       #tempInternalError := MOVE_BLK_VARIANT(SRC := #initialValue,
                                              COUNT := 1,
                                              SRC_INDEX := 0,
                                              DEST_INDEX := #tempSizeCounter,
                                              DEST => #buffer);
     END_FOR;
     IF (#tempInternalError <> #NO_INTERNAL_ERROR) THEN
       #error := true;
       #statusID := #ERROR_MOVE_BLK_VARIANT;
       #status := INT_TO_WORD(#tempInternalError);
     END_IF;
     RETURN;
   END_IF;

   //-----------Program code execution, depending on the Mode parameter-------------
   // The execution of the instructions depends on the signal state of the Mode parameter.

   IF #mode = #NEXT_TASK_TO_EXECUTE THEN


     // If the Mode parameter has the signal state "0",
     // the first entry from the passed ring buffer is returned.

     //this program code section checks whether the ring #buffer is empty.
     //IF this is the CASE, program execution is terminated at this point
     //AND the error code "8001" is output. *)

     IF (#statFirstItemIndex = #BUFFER_IS_EMPTY) THEN
       #error := true;
       #statusID := #ERROR_IN_THIS_BLOCK;
       #status := #BUFFER_EMPTY;
       RETURN;
     END_IF;


     // This program code section returns the first entry of the ring buffer.

     #tempInternalError := MOVE_BLK_VARIANT(SRC := #buffer,
                                            COUNT := 1,
                                            SRC_INDEX := #statFirstItemIndex,
                                            DEST_INDEX := 0,
                                            DEST => #item);

     IF (#tempInternalError = #BUFFER_CONTAINS_ARRAY) THEN

       //This program code section checks whether the ring #buffer contains ARRAY elements.
       //IF it does, the first entry is passed further on
       //AND the index is incremented BY 1. *)

       #tempInternalError := MOVE_BLK_VARIANT(SRC := #initialValue,
                                              COUNT := 1,
                                              SRC_INDEX := 0,
                                              DEST_INDEX := #statFirstItemIndex,
                                              DEST => #buffer);

       // This program code section calculates the new index of the first entry.

       #tempNewFirstItemIndex := #statFirstItemIndex + 1;
       #tempNewFirstItemIndex := #tempNewFirstItemIndex MOD UDINT_TO_INT(#tempPufferSize);

       // This program section checks whether the ring buffer is empty.        
       IF (#statNextEmptyItemIndex = #tempNewFirstItemIndex) THEN
         // If the ring buffer is empty, the index is set to 0.            
         #statFirstItemIndex := -1;
         #statNextEmptyItemIndex := 0;
       ELSE
         // The index of the first entry is changed.            
         #statFirstItemIndex := #tempNewFirstItemIndex;
       END_IF;
     END_IF;
   ELSE

     // If the Mode parameter has the signal state "1", the entry is written to the passed ring buffer.

     //this program code section checks whether the ring #buffer is full.
     //IF this is the CASE, program execution is terminated at this point
     //AND the error code "8002" is output. *)

     IF (#statNextEmptyItemIndex = #statFirstItemIndex) THEN
       #error := true;
       #statusID := #ERROR_IN_THIS_BLOCK;
       #status := #BUFFER_FULL;
       RETURN;
     END_IF;

     // This program code section writes the entry to the ring buffer.   
     #tempInternalError := MOVE_BLK_VARIANT(SRC := #item,
                                            COUNT := 1,
                                            SRC_INDEX := 0,
                                            DEST_INDEX := #statNextEmptyItemIndex,
                                            DEST => #buffer);

     IF (#tempInternalError = #NO_INTERNAL_ERROR) THEN

       // This program code section increments the index by 1 and calculates the new empty entry index.        
       #tempNewNextEmptyItemIndex := #statNextEmptyItemIndex + 1;
       #tempNewNextEmptyItemIndex := #tempNewNextEmptyItemIndex MOD UDINT_TO_INT(#tempPufferSize);
       #statNextEmptyItemIndex := #tempNewNextEmptyItemIndex;

       //This program code section checks which index the "#firstItemIndex" tag has.
       //IF the number = -1, the ring buffer is initialized
       //AND the entry is written TO the ring #buffer.
       //Therefore, "0" must be assigned TO the tag.

       IF (#statFirstItemIndex = #BUFFER_INITIALIZED) THEN
         #statFirstItemIndex := 0;
       END_IF;
     END_IF;
   END_IF;

   //-------------------------Local error handling----------------------------
   //This program code section checks whether a "Local" #error has occurred.
   //IF This is the CASE, program execution is terminated at This point
   //AND the error code of MOV_BLK_VARIANT is output. *)

   IF (#tempInternalError <> #NO_INTERNAL_ERROR) THEN
     #error := true;
     #statusID := #ERROR_MOVE_BLK_VARIANT;
     #status := INT_TO_WORD(#tempInternalError);
     RETURN;
   END_IF;

   #status := #NO_ERROR;
END_FUNCTION_BLOCK

FUNCTION_BLOCK "LGF_ShellSortInt"   // FB10018, SCL
{ S7_Optimized_Access := 'TRUE' }
   VAR_INPUT
      mode : Bool;   // FALSE: Sort ascending; TRUE: Sort descending
   END_VAR
   VAR_OUTPUT
      error : Bool;   // Error
      statusID : UInt;   // Status ID
      status : Word;   // Status information
   END_VAR
   VAR_IN_OUT
      variantArray : Variant;   // Array to be sorted
   END_VAR
   VAR_TEMP
      tempArrayInt : Array[1..#MAX_ARRAY_ELEMENTS] of Int;   // -
      tempElementCount : Int;   // -
      tempElementCopyCount : UDInt;   // -
      tempMoveBlkError : Int;   // -
      tempIncrement : Int;   // -
      tempForCounter : Int;   // -
      tempExchangeIndex : Int;   // -
      tempExchangeVariable : Int;   // -
      tempTypeTag : Int;   // -
   END_VAR
   VAR CONSTANT
      MAX_ARRAY_ELEMENTS : Int := 1000;   // Max array elements allowed
      NO_ERROR : Word := 16#0000;   // No errors
      NO_CURRENT_JOBS : Word := 16#7000;   // Initial value
      EMPTY_ARRAY : Word := 16#8200;   // Array is empty
      NOT_AN_ARRAY : Word := 16#8201;   // Data type is not an Array
      WRONG_ELEMENT_TYPE : Word := 16#8202;   // Wrong data type of Array element
      TOO_MANY_ELEMENTS : Word := 16#8203;   // Too many Array elements
      ERROR_IN_THIS_BLOCK : UInt := 1;   // Error in this block
      ERROR_MOVE_BLK_VARIANT_R : UInt := 2;   // Error/status of subordinate block "MOVE_BLK_VARIANT" when reading
      ERROR_MOVE_BLK_VARIANT_W : UInt := 3;   // Error/status of subordinate block "MOVE_BLK_VARIANT" when writing
   END_VAR
BEGIN
   //=============================================================================
   // SIEMENS AG
   // (c)Copyright 2017
   //-----------------------------------------------------------------------------
   // Library:       LGF (Library General Functions)
   // Tested with:   CPU1212C DC/DC/DC FW:V4.2
   // Engineering:   TIA Portal V14 Update 1
   // Restrictions:  -
   // Requirements:  PLC (S7-1200 / S7-1500)
   // Functionality: A shellsort algorithm with a complexity between 'n^2' and
   //                'n log n' for average, best and worst case inputs and space
   //                complexity '1'.
   //                The block accepts an Integer array as an inOut-variable and
   //                returns the sorted version of the array in the same variable
   //-----------------------------------------------------------------------------
   // Change log table:
   // Version  Date        Expert in charge / Changes applied
   // 01.00.00 19.08.2015  Siemens Industry Online Support
   //                      First released version
   // 01.01.00 19.05.2016  Siemens Industry Online Support
   //                      New function: reverse sort
   // 01.01.01 02.01.2017  Siemens Industry Online Support
   //                      Upgrade: TIA Portal V14 Update 1
   // 01.01.02 17.08.2018  Siemens Industry Online Support
   //                      Upgrade: TIA V15 Update 2
   // 01.01.03 23.11.2018  Siemens Industry Online Support
   //                      Upgrade: TIA V15.1
   // 02.00.00 29.01.2019  Siemens Industry Online Support
   //                      Output "done" removed (not necessary, because only one cycle)
   //-----------------------------------------------------------------------------
   //Status Codes:
   // 16#7000:  No current jobs
   // 16#0000:  Job finished; Note: There is no "Busy"-Status because the block is
   //           finished within a single cycle
   // 16#8200:  Error: Parameter is an an array with only one element
   // 16#8201:  Error: Parameter is not an array
   // 16#8202:  Error: Parameter is an array of the wrong type
   //           (correct type is Integer)
   // 16#8203:  Error: There are too many Elements in the array
   //          (default: max. 1000 Elements)
   //=============================================================================

   // Change note: If you wish to use this shellsort block for other datatypes,
   // you simply need to change the following variables to that type
   // 1. tempExchangeVariable
   // 2. tempTypeTag
   // 3. tempArray<Type>
   // Space note: If you wish to reduce the space of this block, you may reduce the
   // size OF the tempArray<Type> TO one just big enough FOR your specific purpose
   // It is not recommended to increase the size significantly.

   // Initialization
   #tempElementCount := 0;
   #tempElementCopyCount := 0;
   #tempMoveBlkError := 0;
   #tempIncrement := 0;
   #tempForCounter := 0;
   #tempExchangeIndex := 0;
   #tempExchangeVariable := 0;
   #tempTypeTag := 0;

   // Set "No current job" status
   #error := false;
   #statusID := #ERROR_IN_THIS_BLOCK;
   #status := #NO_CURRENT_JOBS;


   // If the variant inOut-parameter is not an array, set error status 8201
   IF (IS_ARRAY(#variantArray) = false) THEN
     #error := true;
     #statusID := #ERROR_IN_THIS_BLOCK;
     #status := #NOT_AN_ARRAY;
     RETURN;
   ELSE
     IF TypeOfElements(#variantArray) = TypeOf(#tempTypeTag) THEN
       // If the parameter is an array of the type integer, get the element count
       #tempElementCopyCount := CountOfElements(#variantArray);
       #tempElementCount := UDINT_TO_INT(CountOfElements(#variantArray));
       // Check whether the variant array contains less than the maximum possible amount of elements
       IF #tempElementCount > #MAX_ARRAY_ELEMENTS THEN
         #error := true;
         #statusID := #ERROR_IN_THIS_BLOCK;
         #status := #TOO_MANY_ELEMENTS;
         RETURN;
       END_IF;
     ELSE
       // If the parameter is an array but not of the type integer, set an error status
       #error := true;
       #statusID := #ERROR_IN_THIS_BLOCK;
       #status := #WRONG_ELEMENT_TYPE;
       RETURN;
     END_IF;
   END_IF;

   // If there are more than zero elements to sort, begin sorting    
   IF #tempElementCount > 1 AND #error = false THEN

     // Read the elements of the incoming variant-array and write into the local array
     #tempMoveBlkError := MOVE_BLK_VARIANT(COUNT := #tempElementCopyCount,
                                           DEST => #tempArrayInt,
                                           DEST_INDEX := 0,
                                           SRC := #variantArray,
                                           SRC_INDEX := 0);

     // Error handling for MOVE_BLK_VARIANT
     IF #tempMoveBlkError <> 0 THEN
       #error := true;
       #statusID := #ERROR_MOVE_BLK_VARIANT_R;
       #status := INT_TO_WORD(#tempMoveBlkError);
       RETURN;
     END_IF;

     // ShellSort Start
     #tempIncrement := 1;
     REPEAT
       #tempIncrement := (3 * #tempIncrement) + 1;
     UNTIL #tempIncrement > #tempElementCount
     END_REPEAT;

     REPEAT
       #tempIncrement := DINT_TO_INT(TRUNC(#tempIncrement / 3));
       FOR #tempForCounter := (#tempIncrement + 1) TO #tempElementCount DO
         #tempExchangeVariable := #tempArrayInt[#tempForCounter];
         #tempExchangeIndex := #tempForCounter;

         IF #mode  // Modification Version 02.00.00
         THEN      //mode = TRUE --> sort descending  
           WHILE ((#tempArrayInt[#tempExchangeIndex - #tempIncrement] < #tempExchangeVariable)) DO
             #tempArrayInt[#tempExchangeIndex] := #tempArrayInt[#tempExchangeIndex - #tempIncrement];
             #tempExchangeIndex := #tempExchangeIndex - #tempIncrement;
             IF (#tempExchangeIndex <= #tempIncrement) THEN
               GOTO EXITWhile;
             END_IF;
           END_WHILE;
         ELSE      // mode = FALSE --> sort ascending
           WHILE ((#tempArrayInt[#tempExchangeIndex - #tempIncrement] > #tempExchangeVariable)) DO
             #tempArrayInt[#tempExchangeIndex] := #tempArrayInt[#tempExchangeIndex - #tempIncrement];
             #tempExchangeIndex := #tempExchangeIndex - #tempIncrement;
             IF (#tempExchangeIndex <= #tempIncrement) THEN
               GOTO EXITWhile;
             END_IF;
           END_WHILE;
         END_IF;

       EXITWhile:
         #tempArrayInt[#tempExchangeIndex] := #tempExchangeVariable;
       END_FOR;
     UNTIL #tempIncrement <= 1
     END_REPEAT;
     // ShellSort End

     // Write the elements of the local array back to the variant array
     #tempMoveBlkError := MOVE_BLK_VARIANT(COUNT := #tempElementCopyCount,
                                           DEST => #variantArray,
                                           DEST_INDEX := 0,
                                           SRC := #tempArrayInt,
                                           SRC_INDEX := 0);

     // Error handling for MOVE_BLK_VARIANT
     IF #tempMoveBlkError <> 0 THEN
       #statusID := #ERROR_MOVE_BLK_VARIANT_W;
       #status := INT_TO_WORD(#tempMoveBlkError);
       RETURN;
     END_IF;

     // Set output status 
     #status := #NO_ERROR;

   ELSIF #tempElementCount <= 1 THEN
     // If there are 0 elements in the array, set status to "Error: Parameter is an empty array"
     #error := true;
     #statusID := #ERROR_IN_THIS_BLOCK;
     #status := #EMPTY_ARRAY;
   END_IF;
END_FUNCTION_BLOCK

FUNCTION_BLOCK "LGF_ShellSortReal"   // FB10019, SCL
{ S7_Optimized_Access := 'TRUE' }
   VAR_INPUT
      mode : Bool;   // FALSE: Sort ascending; TRUE: Sort descending
   END_VAR
   VAR_OUTPUT
      error : Bool;   // Error
      statusID : UInt;   // Status ID
      status : Word;   // Status information
   END_VAR
   VAR_IN_OUT
      variantArray : Variant;   // Array to be sorted
   END_VAR
   VAR_TEMP
      tempArrayReal : Array[1..#MAX_ARRAY_ELEMENTS] of Real;   // -
      tempElementCount : Int;   // -
      tempElementCopyCount : UDInt;   // -
      tempMoveBlkError : Int;   // -
      tempIncrement : Int;   // -
      tempForCounter : Int;   // -
      tempExchangeIndex : Int;   // -
      tempExchangeVariable : Real;   // -
      tempTypeTag : Real;   // -
   END_VAR
   VAR CONSTANT
      MAX_ARRAY_ELEMENTS : Int := 1000;   // Max array elements allowed
      NO_ERROR : Word := 16#0000;   // No errors
      NO_CURRENT_JOBS : Word := 16#7000;   // Initial value
      EMPTY_ARRAY : Word := 16#8200;   // Array is empty
      NOT_AN_ARRAY : Word := 16#8201;   // Data type is not an Array
      WRONG_ELEMENT_TYPE : Word := 16#8202;   // Wrong data type of Array element
      TOO_MANY_ELEMENTS : Word := 16#8203;   // Too many Array elements
      ERROR_IN_THIS_BLOCK : UInt := 1;   // Error in this block
      ERROR_MOVE_BLK_VARIANT_R : UInt := 2;   // Error/status of subordinate block "MOVE_BLK_VARIANT" when reading
      ERROR_MOVE_BLK_VARIANT_W : UInt := 3;   // Error/status of subordinate block "MOVE_BLK_VARIANT" when writing
   END_VAR
BEGIN
   //=============================================================================
   // SIEMENS AG
   // (c)Copyright 2017
   //-----------------------------------------------------------------------------
   // Library:       LGF (Library General Functions)
   // Tested with:   CPU1212C DC/DC/DC FW:V4.2
   // Engineering:   TIA Portal V14 Update 1
   // Restrictions:  -
   // Requirements:  PLC (S7-1200 / S7-1500)
   // Functionality: A shellsort algorithm with a complexity between 'n^2' and
   //                'n log n' for average, best and worst case inputs and space
   //                complexity '1'.
   //                The block accepts a Real array as an inOut-variable and
   //                returns the sorted version of the array in the same variable
   //-----------------------------------------------------------------------------
   // Change log table:
   // Version  Date        Expert in charge / Changes applied
   // 01.00.00 19.08.2015  Siemens Industry Online Support
   //                      First released version
   // 01.01.00 19.05.2016  Siemens Industry Online Support
   //                      New function: reverse sort
   // 01.01.01 02.01.2017  Siemens Industry Online Support
   //                      Upgrade: TIA Portal V14 Update 1
   // 01.01.02 17.08.2018  Siemens Industry Online Support
   //                      Upgrade: TIA V15 Update 2
   // 01.01.03 23.11.2018  Siemens Industry Online Support
   //                      Upgrade: TIA V15.1
   // 02.00.00 29.01.2019  Siemens Industry Online Support
   //                      Output "done" removed (not necessary, because only one cycle)
   //-----------------------------------------------------------------------------
   //Status Codes:
   // 16#7000:  No current jobs
   // 16#0000:  Job finished; Note: There is no "Busy"-Status because the block is
   //           finished within a single cycle
   // 16#8200:  Error: Parameter is an array with only one element
   // 16#8201:  Error: Parameter is not an array
   // 16#8202:  Error: Parameter is an array of the wrong type
   //           (correct type is Real)
   // 16#8203:  Error: There are too many Elements in the array
   //           (default: max. 1000 Elements)
   //=============================================================================

   // Change note: If you wish to use this shellsort block for other datatypes,
   // you simply need to change the following variables to that type
   // 1. tempExchangeVariable
   // 2. tempTypeTag
   // 3. tempArray<Type>
   // Space note: If you wish to reduce the space of this block, you may reduce the
   // size of the tempArray<Type> to one just big enough for your specific purpose
   // It is not recommended to increase the size significantly.

   // Initialization
   #tempElementCount := 0;
   #tempElementCopyCount := 0;
   #tempMoveBlkError := 0;
   #tempIncrement := 0;
   #tempForCounter := 0;
   #tempExchangeIndex := 0;
   #tempExchangeVariable := 0;
   #tempTypeTag := 0;

   // Set "No current job" status
   #error := false;
   #statusID := #ERROR_IN_THIS_BLOCK;
   #status := #NO_CURRENT_JOBS;


   // If the variant inOut-parameter is not an array, set error status 8201
   IF (IS_ARRAY(#variantArray) = false) THEN
     #error := true;
     #statusID := #ERROR_IN_THIS_BLOCK;
     #status := #NOT_AN_ARRAY;
     RETURN;
   ELSE
     IF TypeOfElements(#variantArray) = TypeOf(#tempTypeTag) THEN
       // If the parameter is an array of the type real, get the element count
       #tempElementCopyCount := CountOfElements(#variantArray);
       #tempElementCount := UDINT_TO_INT(CountOfElements(#variantArray));
       // Check whether the variant array contains less than the maximum possible amount of elements
       IF #tempElementCount > #MAX_ARRAY_ELEMENTS THEN
         #error := true;
         #statusID := #ERROR_IN_THIS_BLOCK;
         #status := #TOO_MANY_ELEMENTS;
         RETURN;
       END_IF;
     ELSE
       // If the parameter is an array but not of the type real, set an error status
       #error := true;
       #statusID := #ERROR_IN_THIS_BLOCK;
       #status := #WRONG_ELEMENT_TYPE;
       RETURN;
     END_IF;
   END_IF;

   // If there are more than zero elements to sort, begin sorting    
   IF #tempElementCount > 1 AND #error = false THEN

     // Read the elements of the incoming variant-array and write into the local array
     #tempMoveBlkError := MOVE_BLK_VARIANT(COUNT := #tempElementCopyCount,
                                           DEST => #tempArrayReal,
                                           DEST_INDEX := 0,
                                           SRC := #variantArray,
                                           SRC_INDEX := 0);

     // Error handling for MOVE_BLK_VARIANT
     IF #tempMoveBlkError <> 0 THEN
       #error := true;
       #statusID := #ERROR_MOVE_BLK_VARIANT_R;
       #status := INT_TO_WORD(#tempMoveBlkError);
       RETURN;
     END_IF;

     // ShellSort Start
     #tempIncrement := 1;
     REPEAT
       #tempIncrement := (3 * #tempIncrement) + 1;
     UNTIL #tempIncrement > #tempElementCount
     END_REPEAT;

     REPEAT
       #tempIncrement := DINT_TO_INT(TRUNC(#tempIncrement / 3));
       FOR #tempForCounter := (#tempIncrement + 1) TO #tempElementCount DO
         #tempExchangeVariable := #tempArrayReal[#tempForCounter];
         #tempExchangeIndex := #tempForCounter;

         IF #mode  // Modification Version 02.00.00
         THEN      //mode = TRUE --> sort descending  
           WHILE ((#tempArrayReal[#tempExchangeIndex - #tempIncrement] < #tempExchangeVariable)) DO
             #tempArrayReal[#tempExchangeIndex] := #tempArrayReal[#tempExchangeIndex - #tempIncrement];
             #tempExchangeIndex := #tempExchangeIndex - #tempIncrement;
             IF (#tempExchangeIndex <= #tempIncrement) THEN
               GOTO EXITWhile;
             END_IF;
           END_WHILE;
         ELSE      // mode = FALSE --> sort ascending
           WHILE ((#tempArrayReal[#tempExchangeIndex - #tempIncrement] > #tempExchangeVariable)) DO
             #tempArrayReal[#tempExchangeIndex] := #tempArrayReal[#tempExchangeIndex - #tempIncrement];
             #tempExchangeIndex := #tempExchangeIndex - #tempIncrement;
             IF (#tempExchangeIndex <= #tempIncrement) THEN
               GOTO EXITWhile;
             END_IF;
           END_WHILE;
         END_IF;

       EXITWhile:
         #tempArrayReal[#tempExchangeIndex] := #tempExchangeVariable;
       END_FOR;
     UNTIL #tempIncrement <= 1
     END_REPEAT;
     // ShellSort End

     // Write the elements of the local array back to the variant array
     #tempMoveBlkError := MOVE_BLK_VARIANT(COUNT := #tempElementCopyCount,
                                           DEST => #variantArray,
                                           DEST_INDEX := 0,
                                           SRC := #tempArrayReal,
                                           SRC_INDEX := 0);

     // Error handling for MOVE_BLK_VARIANT
     IF #tempMoveBlkError <> 0 THEN
       #statusID := #ERROR_MOVE_BLK_VARIANT_W;
       #status := INT_TO_WORD(#tempMoveBlkError);
       RETURN;
     END_IF;

     // Set output status 
     #status := #NO_ERROR;

   ELSIF #tempElementCount <= 1 THEN
     // If there are 0 elements in the array, set status to "Error: Parameter is an empty array"
     #error := true;
     #statusID := #ERROR_IN_THIS_BLOCK;
     #status := #EMPTY_ARRAY;
   END_IF;
END_FUNCTION_BLOCK

FUNCTION_BLOCK "LGF_ShellSortUInt"   // FB10020, SCL
{ S7_Optimized_Access := 'TRUE' }
   VAR_INPUT
      mode : Bool;   // FALSE: Sort ascending; TRUE: Sort descending
   END_VAR
   VAR_OUTPUT
      error : Bool;   // Error
      statusID : UInt;   // Status ID
      status : Word;   // Status information
   END_VAR
   VAR_IN_OUT
      variantArray : Variant;   // Array to be sorted
   END_VAR
   VAR_TEMP
      tempArrayUInt : Array[1..#MAX_ARRAY_ELEMENTS] of UInt;   // -
      tempElementCount : Int;   // -
      tempElementCopyCount : UDInt;   // -
      tempMoveBlkError : Int;   // -
      tempIncrement : Int;   // -
      tempForCounter : Int;   // -
      tempExchangeIndex : Int;   // -
      tempExchangeVariable : UInt;   // -
      tempTypeTag : UInt;   // -
   END_VAR
   VAR CONSTANT
      MAX_ARRAY_ELEMENTS : Int := 1000;   // Max array elements allowed
      NO_ERROR : Word := 16#0000;   // No errors
      NO_CURRENT_JOBS : Word := 16#7000;   // Initial value
      EMPTY_ARRAY : Word := 16#8200;   // Array is empty
      NOT_AN_ARRAY : Word := 16#8201;   // Data type is not an Array
      WRONG_ELEMENT_TYPE : Word := 16#8202;   // Wrong data type of Array element
      TOO_MANY_ELEMENTS : Word := 16#8203;   // Too many Array elements
      ERROR_IN_THIS_BLOCK : UInt := 1;   // Error in this block
      ERROR_MOVE_BLK_VARIANT_R : UInt := 2;   // Error/status of subordinate block "MOVE_BLK_VARIANT" when reading
      ERROR_MOVE_BLK_VARIANT_W : UInt := 3;   // Error/status of subordinate block "MOVE_BLK_VARIANT" when writing
   END_VAR
BEGIN
   //=============================================================================
   // SIEMENS AG
   // (c)Copyright 2017
   //-----------------------------------------------------------------------------
   // Library:       LGF (Library General Functions)
   // Tested with:   CPU1212C DC/DC/DC FW:V4.2
   // Engineering:   TIA Portal V14
   // Restrictions:  -
   // Requirements:  PLC (S7-1200 / S7-1500)
   // Functionality: A shellsort algorithm with a complexity between 'n^2' and
   //                'n log n' for average, best and worst case inputs and space
   //                complexity '1'.
   //                The block accepts an unsigned Integer array as an
   //                inOut-variable and returns the sorted version of the array in
   //                the same variable
   //-----------------------------------------------------------------------------
   // Change log table:
   // Version  Date        Expert in charge / Changes applied
   // 01.00.00 19.08.2015  Siemens Industry Online Support
   //                      First released version
   // 01.01.00 19.05.2016  Siemens Industry Online Support
   //                      New function: reverse sort
   // 01.01.01 02.01.2017  Siemens Industry Online Support
   //                      Upgrade: TIA Portal V14 Update 1
   // 01.01.02 17.08.2018  Siemens Industry Online Support
   //                      Upgrade: TIA V15 Update 2
   // 01.01.03 23.11.2018  Siemens Industry Online Support
   //                      Upgrade: TIA V15.1
   // 02.00.00 29.01.2019  Siemens Industry Online Support
   //                      Output "done" removed (not necessary, because only one cycle)
   //-----------------------------------------------------------------------------
   //Status Codes:
   // 16#7000:  No current jobs
   // 16#0000:  Job finished     //Note: There is no "Busy"-Status because the
   //           block is finished within a single cycle
   // 16#8200:  Error: Parameter is an array with only one element
   // 16#8201:  Error: Parameter is not an array
   // 16#8202:  Error: Parameter is an array of the wrong type
   //           (correct type is unsigned Integer)
   // 16#8203:  Error: There are too many Elements in the array
   //          (default: max. 1000 Elements)
   //=============================================================================

   // Change note: If you wish to use this shellsort block for other datatypes,
   // you simply need to change the following variables to that type
   // 1. tempExchangeVariable
   // 2. tempTypeTag
   // 3. tempArray<Type>
   // Space note: If you wish to reduce the space of this block, you may reduce the
   // size of the tempArray<Type> to one just big enough for your specific purpose
   // It is not recommended to increase the size significantly.

   // Initialization
   #tempElementCount := 0;
   #tempElementCopyCount := 0;
   #tempMoveBlkError := 0;
   #tempIncrement := 0;
   #tempForCounter := 0;
   #tempExchangeIndex := 0;
   #tempExchangeVariable := 0;
   #tempTypeTag := 0;

   // Set "No current job" status
   #error := false;
   #statusID := #ERROR_IN_THIS_BLOCK;
   #status := #NO_CURRENT_JOBS;


   // If the variant InOut-parameter is not an array, set error status 8201
   IF (IS_ARRAY(#variantArray) = false) THEN
     #error := true;
     #statusID := #ERROR_IN_THIS_BLOCK;
     #status := #NOT_AN_ARRAY;
     RETURN;
   ELSE
     IF TypeOfElements(#variantArray) = TypeOf(#tempTypeTag) THEN
       // If the parameter is an array of the type unsigned integer, get the element count
       #tempElementCopyCount := CountOfElements(#variantArray);
       #tempElementCount := UDINT_TO_INT(CountOfElements(#variantArray));
       // Check whether the variant array contains less than the maximum possible amount of elements
       IF #tempElementCount > #MAX_ARRAY_ELEMENTS THEN
         #error := true;
         #statusID := #ERROR_IN_THIS_BLOCK;
         #status := #TOO_MANY_ELEMENTS;
         RETURN;
       END_IF;
     ELSE
       //If the parameter is an array but not of the type unsigned integer, set an error status
       #error := true;
       #statusID := #ERROR_IN_THIS_BLOCK;
       #status := #WRONG_ELEMENT_TYPE;
       RETURN;
     END_IF;
   END_IF;

   //If there are more than zero elements to sort, begin sorting    
   IF #tempElementCount > 1 AND #error = false THEN

     //Read the elements of the incoming variant-array and write into the local array
     #tempMoveBlkError := MOVE_BLK_VARIANT(COUNT := #tempElementCopyCount,
                                           DEST => #tempArrayUInt,
                                           DEST_INDEX := 0,
                                           SRC := #variantArray,
                                           SRC_INDEX := 0);

     // Error handling for MOVE_BLK_VARIANT
     IF #tempMoveBlkError <> 0 THEN
       #error := true;
       #statusID := #ERROR_MOVE_BLK_VARIANT_R;
       #status := INT_TO_WORD(#tempMoveBlkError);
       RETURN;
     END_IF;

     // ShellSort Start
     #tempIncrement := 1;
     REPEAT
       #tempIncrement := (3 * #tempIncrement) + 1;
     UNTIL #tempIncrement > #tempElementCount
     END_REPEAT;

     REPEAT
       #tempIncrement := DINT_TO_INT(TRUNC(#tempIncrement / 3));
       FOR #tempForCounter := (#tempIncrement + 1) TO #tempElementCount DO
         #tempExchangeVariable := #tempArrayUInt[#tempForCounter];
         #tempExchangeIndex := #tempForCounter;

         IF #mode  // Modification Version 02.00.00
         THEN      //mode = TRUE --> sort descending  
           WHILE ((#tempArrayUInt[#tempExchangeIndex - #tempIncrement] < #tempExchangeVariable)) DO
             #tempArrayUInt[#tempExchangeIndex] := #tempArrayUInt[#tempExchangeIndex - #tempIncrement];
             #tempExchangeIndex := #tempExchangeIndex - #tempIncrement;
             IF (#tempExchangeIndex <= #tempIncrement) THEN
               GOTO EXITWhile;
             END_IF;
           END_WHILE;
         ELSE      // mode = FALSE --> sort ascending
           WHILE ((#tempArrayUInt[#tempExchangeIndex - #tempIncrement] > #tempExchangeVariable)) DO
             #tempArrayUInt[#tempExchangeIndex] := #tempArrayUInt[#tempExchangeIndex - #tempIncrement];
             #tempExchangeIndex := #tempExchangeIndex - #tempIncrement;
             IF (#tempExchangeIndex <= #tempIncrement) THEN
               GOTO EXITWhile;
             END_IF;
           END_WHILE;
         END_IF;

       EXITWhile:
         #tempArrayUInt[#tempExchangeIndex] := #tempExchangeVariable;
       END_FOR;
     UNTIL #tempIncrement <= 1
     END_REPEAT;
     // ShellSort End

     // Write the elements of the local array back to the variant array
     #tempMoveBlkError := MOVE_BLK_VARIANT(COUNT := #tempElementCopyCount,
                                           DEST => #variantArray,
                                           DEST_INDEX := 0,
                                           SRC := #tempArrayUInt,
                                           SRC_INDEX := 0);

     // Error handling for MOVE_BLK_VARIANT
     IF #tempMoveBlkError <> 0 THEN
       #statusID := #ERROR_MOVE_BLK_VARIANT_W;
       #status := INT_TO_WORD(#tempMoveBlkError);
       RETURN;
     END_IF;

     // Set output status
     #status := #NO_ERROR;

   ELSIF #tempElementCount <= 1 THEN
     // If there are 0 elements in the array, set status to "Error: Parameter is an empty array"
     #error := true;
     #statusID := #ERROR_IN_THIS_BLOCK;
     #status := #EMPTY_ARRAY;
   END_IF;
END_FUNCTION_BLOCK

FUNCTION_BLOCK "LGF_LIFO"   // FB10021, SCL
{ S7_Optimized_Access := 'TRUE' }
   VAR_INPUT
      execute : Bool;   // The instruction is executed when a positive signal edge is detected at the "request" parameter.
      mode : Bool;   // 0 = The first entry in the ring buffer is returned. 1 = An entry is written at the last position in the ring buffer.
      initialValue : Variant;   // Value with which the ARRAY of the ring buffer is initialized.
      resetBuffer : Bool;   // Clearing and initializing the buffer
   END_VAR
   VAR_OUTPUT
      error : Bool;   // Error
      statusID : UInt;   // Status ID
      status : Word;   // Status information
   END_VAR
   VAR_IN_OUT
      item : Variant;   // The entry that is either returned from the ring buffer or written to the ring buffer
      buffer : Variant;   // An ARRAY that is used as a ring buffer.
   END_VAR
   VAR
      statEdgeUpm : Bool;   // Edge memory bit in which the RLO of the previous query is saved.
      statLastItemIndex : Int := -1;   // Index of the newest entry in the ring buffer
      statNextEmptyItemIndex : Int := 0;   // Index of the next free entry in the ring buffer
   END_VAR
   VAR_TEMP
      tempInternalError : Int;   // Error information
      tempPufferSize : UDInt;   // Number of ARRAY elements in the ring buffer
      tempSizeCounter : Int;   // Size counter
   END_VAR
   VAR CONSTANT
      NO_ERROR : Word := 16#0000;   // No errors
      NO_CURRENT_JOBS : Word := 16#7000;   // Initial value
      BUFFER_EMPTY : Word := 16#8001;   // The buffer is empty
      BUFFER_FULL : Word := 16#8002;   // The buffer is full
      NO_ARRAY : Word := 16#8200;   // No array is present at the input "buffer"
      WRONG_TYPE_1 : Word := 16#8201;   // The data type of the InOut parameter "item" does not correspond to the data type of the array elements of the input "buffer"
      WRONG_TYPE_2 : Word := 16#8202;   // The data type of the input "initialValue" does not correspond to the data type of the InOut parameter "item"
      ERROR_IN_THIS_BLOCK : UInt := 1;   // Error in this block
      ERROR_MOVE_BLK_VARIANT : UInt := 2;   // Error/status of subordinate block "MOVE_BLK_VARIANT"
      NEXT_TASK_TO_EXECUTE : Bool := false;   // Next task to execute
      BUFFER_IS_EMPTY : Int := -1;   // Buffer is empty
      BUFFER_CONTAINS_ARRAY : Int := 0;   // Buffer contains array
      NO_INTERNAL_ERROR : Int := 0;   // No internal error
      BUFFER_INITIALIZED : Int := -1;   // Buffer initialized
      RESET : Bool := true;   // Reset
   END_VAR
BEGIN
   //=============================================================================
   // SIEMENS AG
   // (c)Copyright 2017
   //-----------------------------------------------------------------------------
   // Library:       LGF (Library General Functions)
   // Tested with:   CPU1212C DC/DC/DC FW:V4.2
   // Engineering:   TIA Portal V14
   // Restrictions:  -
   // Requirements:  PLC (S7-1200 / S7-1500)
   // Functionality: LIFO(Last In First Out)-functionblock
   //-----------------------------------------------------------------------------
   // Change log table:
   // Version  Date        Expert in charge / Changes applied
   // 01.00.00 10.07.2018  Siemens Industry Online Support
   //                      First released version
   // 01.00.01 17.08.2018  Siemens Industry Online Support
   //                      Upgrade: TIA V15 Update 2
   // 01.00.02 23.11.2018  Siemens Industry Online Support
   //                      Upgrade: TIA V15.1
   // 02.00.00 29.01.2019  Siemens Industry Online Support
   //                      Output "done" removed (not necessary, because only one cycle)
   //=============================================================================

   //This program code section is only executed once after a negative signal edge.
   IF (#execute = FALSE)
     AND (#statEdgeUpm = TRUE)
   THEN
     // If no error occurred during program execution, the error code "0000" is output.  
     #error := FALSE;
     #statusID := #ERROR_IN_THIS_BLOCK;
     #status := #NO_CURRENT_JOBS;
   END_IF;

   //This program code section is only executed once after a positive signal edge.
   //IF there is no change in the signal state OF the result OF logic operation,
   //the program processing OF the "FIFOQueue" FB is terminated.
   //
   IF (#execute <> TRUE)
     OR (#statEdgeUpm <> FALSE)
   THEN
     #statEdgeUpm := #execute;
     RETURN;
   END_IF;
   #statEdgeUpm := #execute;

   // ------Validation of whether all parameter inputs are valid.----

   //This program code section checks whether the ring #buffer is an ARRAY.
   //IF so, the number OF the ARRAY elements is read out.
   //IF it is NOT an ARRAY, the program execution is terminated at this point
   //AND the status code "8200" is output.

   IF (NOT (IS_ARRAY(#buffer)))
   THEN
     #error := TRUE;
     #statusID := #ERROR_IN_THIS_BLOCK;
     #status := #NO_ARRAY;
     RETURN;
   ELSE
     #tempPufferSize := CountOfElements(#buffer);
   END_IF;

   //This program code section checks whether the data type OF the ARRAY elements matches
   //the data type OF the entry (tag #item). IF the data types DO NOT match,
   //the program execution is terminated at this point AND the error code "8201" is output.

   IF (NOT (TypeOf(#item) = TypeOfElements(#buffer)))
   THEN
     #error := TRUE;
     #statusID := #ERROR_IN_THIS_BLOCK;
     #status := #WRONG_TYPE_1;
     RETURN;
   END_IF;

   //This program code section checks whether the initial value OF the ring #buffer
   //matches the entry (tag #item). IF the data types DO NOT match,
   //the program execution is terminated at this point
   //AND the error code "8202" is output. *)

   IF (NOT (TypeOf(#item) = TypeOf(#initialValue)))
   THEN
     #error := TRUE;
     #statusID := #ERROR_IN_THIS_BLOCK;
     #status := #WRONG_TYPE_2;
     RETURN;
   END_IF;

   //If reset is "TRUE" the buffer and their  counters are resetted
   IF (#resetBuffer = #RESET)
   THEN
     #statLastItemIndex := -1;
     #statNextEmptyItemIndex := 0;

     FOR #tempSizeCounter := 0 TO UDINT_TO_INT(#tempPufferSize - 1) DO

       #tempInternalError := MOVE_BLK_VARIANT(SRC := #initialValue,
                                              COUNT := 1,
                                              SRC_INDEX := 0,
                                              DEST_INDEX := #tempSizeCounter,
                                              DEST => #buffer);
     END_FOR;

     IF (#tempInternalError <> #NO_INTERNAL_ERROR)
     THEN
       #error := TRUE;
       #statusID := #ERROR_MOVE_BLK_VARIANT;
       #status := INT_TO_WORD(#tempInternalError);
     END_IF;
     RETURN;
   END_IF;


   //-----------Program code execution, depending on the Mode parameter-------------
   // The execution of the instructions depends on the signal state of the Mode parameter.

   IF (#mode = #NEXT_TASK_TO_EXECUTE)
   THEN
     // If the Mode parameter has the signal state "0",
     // the first entry from the passed ring buffer is returned.

     //this program code section checks whether the ring #buffer is empty.
     //IF this is the CASE, program execution is terminated at this point
     //AND the error code "8001" is output. *)

     IF (#statLastItemIndex = #BUFFER_IS_EMPTY)
     THEN
       #error := TRUE;
       #statusID := #ERROR_IN_THIS_BLOCK;
       #status := #BUFFER_EMPTY;
       RETURN;
     END_IF;

     // This program code section returns the first entry of the ring buffer.
     #tempInternalError := MOVE_BLK_VARIANT(SRC := #buffer,
                                            COUNT := 1,
                                            SRC_INDEX := #statLastItemIndex,
                                            DEST_INDEX := 0,
                                            DEST => #item);

     IF (#tempInternalError = #BUFFER_CONTAINS_ARRAY)
     THEN
       //This program code section checks whether the ring #buffer contains ARRAY elements.
       //IF it does, the first entry is passed further on
       //AND the index is incremented BY 1. *)

       #tempInternalError := MOVE_BLK_VARIANT(SRC := #initialValue,
                                              COUNT := 1,
                                              SRC_INDEX := 0,
                                              DEST_INDEX := #statLastItemIndex,
                                              DEST => #buffer);

       // This program code section decrements the index by 1 for reading and writing.
       #statLastItemIndex := #statLastItemIndex - 1;
       #statNextEmptyItemIndex := #statNextEmptyItemIndex - 1;

     END_IF;

   ELSE
     // If the Mode parameter has the signal state "1", the entry is written to the passed ring buffer.

     //this program code section checks whether the ring #buffer is full.
     //IF this is the CASE, program execution is terminated at this point
     //AND the error code "8002" is output. *)

     IF (#statNextEmptyItemIndex >= #tempPufferSize)
     THEN
       #error := TRUE;
       #statusID := #ERROR_IN_THIS_BLOCK;
       #status := #BUFFER_FULL;
       RETURN;
     END_IF;

     // This program code section writes the entry to the ring buffer.   
     #tempInternalError := MOVE_BLK_VARIANT(SRC := #item,
                                            COUNT := 1,
                                            SRC_INDEX := 0,
                                            DEST_INDEX := #statNextEmptyItemIndex,
                                            DEST => #buffer);

     IF (#tempInternalError = #NO_INTERNAL_ERROR)
     THEN
       // This program code section increments the index by 1 for reading and writing.        
       #statLastItemIndex := #statLastItemIndex + 1;
       #statNextEmptyItemIndex := #statNextEmptyItemIndex + 1;
     END_IF;
   END_IF;

   //-------------------------Local error handling----------------------------
   //This program code section checks whether a "Local" #error has occurred.
   //IF This is the CASE, program execution is terminated at This point
   //AND the error code of MOV_BLK_VARIANT is output. *)

   IF (#tempInternalError <> #NO_INTERNAL_ERROR)
   THEN
     #error := TRUE;
     #statusID := #ERROR_MOVE_BLK_VARIANT;
     #status := INT_TO_WORD(#tempInternalError);
     RETURN;
   END_IF;

   #status := #NO_ERROR;
END_FUNCTION_BLOCK

FUNCTION "LGF_CRC8" : Byte   // FC4, SCL
{ S7_Optimized_Access := 'TRUE' }
VERSION : 0.1
   VAR_INPUT
      initValue : Byte;   // Initial value of CRC
      mask : Byte;   // Mask (CRC polynomial) / generator polynomial
   END_VAR
   VAR_IN_OUT
      inputArray : Array[*] of Byte;   // Input array / data stream
   END_VAR
   VAR_TEMP
      tempCRC : Byte;   // CRC checksum
      tempLowerLimit : DInt;   // Lower limit of input array
      tempUpperLimit : DInt;   // Upper limit of input array
      tempIndex1 : Int;   // -
      tempIndex2 : Int;   // -
   END_VAR
   // Ret_Val : CRC8 checksum
BEGIN
   //=============================================================================
   // Siemens AG
   // (c)Copyright 2017
   //-----------------------------------------------------------------------------
   // Library:       LGF (Library General Functions)
   // Tested with:   CPU1212C DC/DC/DC FW:V4.2
   // Engineering:   TIA Portal V14 SP1 Upd 5
   // Restrictions:  -
   // Requirements:  PLC (S7-1200 / S7-1500)
   // Functionality: CRC8
   //-----------------------------------------------------------------------------
   // Change log table:
   // Version  Date        In charge / Changes applied
   // 01.00.00 03.07.2018  Siemens Industry Online Support
   //                      First released version
   // 01.00.01 17.08.2018  Siemens Industry Online Support
   //                      Upgrade: TIA V15 Update 2
   // 01.00.02 23.11.2018  Siemens Industry Online Support
   //                      Upgrade: TIA V15.1
   //=============================================================================

   #tempLowerLimit := LOWER_BOUND(ARR := #inputArray, DIM := 1);
   #tempUpperLimit := UPPER_BOUND(ARR := #inputArray, DIM := 1);

   #tempCRC := #initValue;

   FOR #tempIndex1 := #tempLowerLimit TO #tempUpperLimit DO

     #tempCRC := #tempCRC XOR #inputArray[#tempIndex1];

     FOR #tempIndex2 := 0 TO 7 DO
       IF ((#tempCRC AND 16#80) <> 0)
       THEN
         #tempCRC := SHL(IN := #tempCRC, N := 1) XOR #mask;
       ELSE
         #tempCRC := SHL(IN := #tempCRC, N := 1);
       END_IF;
     END_FOR;

   END_FOR;

   #LGF_CRC8 := #tempCRC;
END_FUNCTION

FUNCTION "LGF_CRC8For1Byte" : Byte   // FC5, SCL
{ S7_Optimized_Access := 'TRUE' }
VERSION : 0.1
   VAR_INPUT
      initValue : Byte;   // Initial value of CRC
      mask : Byte;   // Mask (CRC polynomial) / generator polynomial
      inputByte : Byte;   // Input value
   END_VAR
   VAR_TEMP
      tempCRC : Byte;   // CRC checksum
      tempIndex : Int;   // -
   END_VAR
   // Ret_Val : CRC checksum
BEGIN
   //=============================================================================
   // Siemens AG
   // (c)Copyright 2017
   //-----------------------------------------------------------------------------
   // Library:       LGF (Library General Functions)
   // Tested with:   CPU1212C DC/DC/DC FW:V4.2
   // Engineering:   TIA Portal V14 SP1 Upd 5
   // Restrictions:  -
   // Requirements:  PLC (S7-1200 / S7-1500)
   // Functionality: CRC8 for 1 byte
   //-----------------------------------------------------------------------------
   // Change log table:
   // Version  Date        In charge / Changes applied
   // 01.00.00 03.07.2018  Siemens Industry Online Support
   //                      First released version
   // 01.00.01 17.08.2018  Siemens Industry Online Support
   //                      Upgrade: TIA V15 Update 2
   // 01.00.02 23.11.2018  Siemens Industry Online Support
   //                      Upgrade: TIA V15.1
   //=============================================================================

   #tempCRC := #initValue XOR #inputByte;

   FOR #tempIndex := 0 TO 7 DO
     IF ((#tempCRC AND 16#80) <> 0)
     THEN
       #tempCRC := SHL(IN := #tempCRC, N := 1) XOR #mask;
     ELSE
       #tempCRC := SHL(IN := #tempCRC, N := 1);
     END_IF;
   END_FOR;

   #LGF_CRC8For1Byte := #tempCRC;
END_FUNCTION

FUNCTION "LGF_CRC16" : Word   // FC6, SCL
{ S7_Optimized_Access := 'TRUE' }
VERSION : 0.1
   VAR_INPUT
      initValue : Word;   // Initial value of CRC
      mask : Word;   // Mask (CRC polynomial) / generator polynomial
   END_VAR
   VAR_IN_OUT
      inputArray : Array[*] of Byte;   // Input array / data stream
   END_VAR
   VAR_TEMP
      tempCRC : Word;   // CRC checksum
      tempLowerLimit : DInt;   // Lower limit of input array
      tempUpperLimit : DInt;   // Upper limit of input array
      tempIndex1 : Int;   // -
      tempIndex2 : Int;   // -
   END_VAR
   // Ret_Val : CRC16 checksum
BEGIN
   //=============================================================================
   // Siemens AG
   // (c)Copyright 2017
   //-----------------------------------------------------------------------------
   // Library:       LGF (Library General Functions)
   // Tested with:   CPU1212C DC/DC/DC FW:V4.2
   // Engineering:   TIA Portal V14 SP1 Upd 5
   // Restrictions:  -
   // Requirements:  PLC (S7-1200 / S7-1500)
   // Functionality: CRC16
   //-----------------------------------------------------------------------------
   // Change log table:
   // Version  Date        In charge / Changes applied
   // 01.00.00 03.07.2018  Siemens Industry Online Support
   //                      First released version
   // 01.00.01 17.08.2018  Siemens Industry Online Support
   //                      Upgrade: TIA V15 Update 2
   // 01.00.02 23.11.2018  Siemens Industry Online Support
   //                      Upgrade: TIA V15.1
   //=============================================================================

   #tempLowerLimit := LOWER_BOUND(ARR := #inputArray, DIM := 1);
   #tempUpperLimit := UPPER_BOUND(ARR := #inputArray, DIM := 1);

   #tempCRC := #initValue;

   FOR #tempIndex1 := #tempLowerLimit TO #tempUpperLimit DO

     #tempCRC := #tempCRC XOR SHL(IN := BYTE_TO_WORD(#inputArray[#tempIndex1]), N := 8);

     FOR #tempIndex2 := 0 TO 7 DO
       IF ((#tempCRC AND 16#8000) <> 0)
       THEN
         #tempCRC := SHL(IN := #tempCRC, N := 1) XOR #mask;
       ELSE
         #tempCRC := SHL(IN := #tempCRC, N := 1);
       END_IF;
     END_FOR;

   END_FOR;

   #LGF_CRC16 := #tempCRC;
END_FUNCTION

FUNCTION "LGF_CRC32" : DWord   // FC7, SCL
{ S7_Optimized_Access := 'TRUE' }